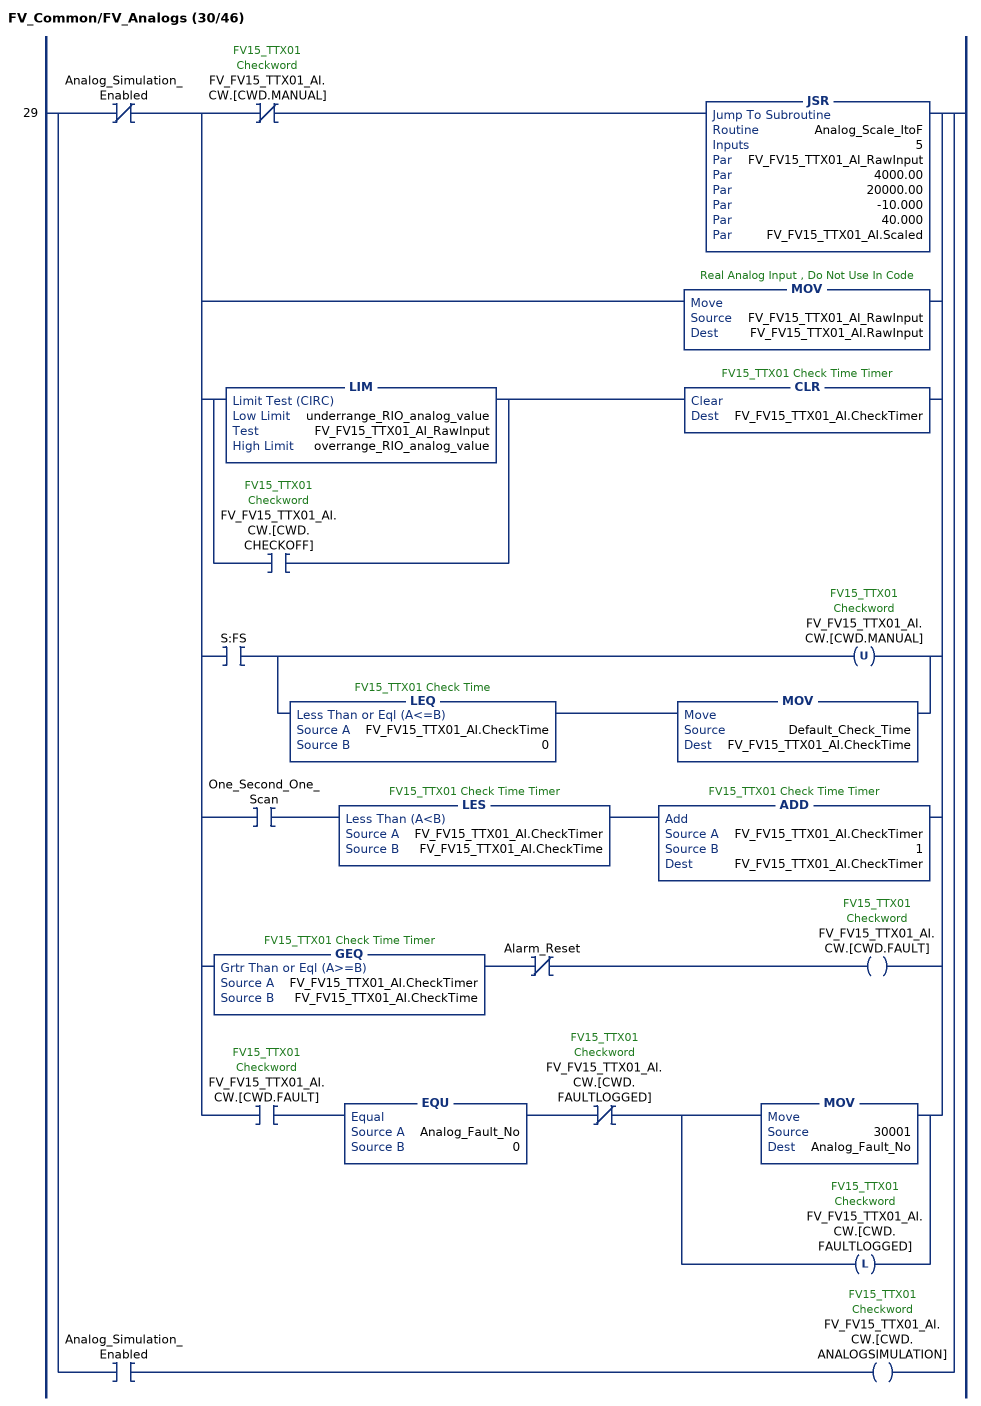
   29: [XIO(Analog_Simulation_Enabled) [XIO(FV_FV15_TTX01_AI.CW.[CWD.MANUAL]) JSR(Analog_Scale_ItoF,5,FV_FV15_TTX01_AI_RawInput,4000.00,20000.00,-10.000,40.000,FV_FV15_TTX01_AI.Scaled) ,MOV(FV_FV15_TTX01_AI_RawInput,FV_FV15_TTX01_AI.RawInput) ,[LIM(underrange_RIO_analog_value,FV_FV15_TTX01_AI_RawInput,overrange_RIO_analog_value) ,XIC(FV_FV15_TTX01_AI.CW.[CWD.CHECKOFF]) ] CLR(FV_FV15_TTX01_AI.CheckTimer) ,XIC(S:FS) [OTU(FV_FV15_TTX01_AI.CW.[CWD.MANUAL]) ,LEQ(FV_FV15_TTX01_AI.CheckTime,0) MOV(Default_Check_Time,FV_FV15_TTX01_AI.CheckTime) ] ,XIC(One_Second_One_Scan) LES(FV_FV15_TTX01_AI.CheckTimer,FV_FV15_TTX01_AI.CheckTime) ADD(FV_FV15_TTX01_AI.CheckTimer,1,FV_FV15_TTX01_AI.CheckTimer) ,GEQ(FV_FV15_TTX01_AI.CheckTimer,FV_FV15_TTX01_AI.CheckTime) XIO(Alarm_Reset) OTE(FV_FV15_TTX01_AI.CW.[CWD.FAULT]) ,XIC(FV_FV15_TTX01_AI.CW.[CWD.FAULT]) EQU(Analog_Fault_No,0) XIO(FV_FV15_TTX01_AI.CW.[CWD.FAULTLOGGED]) [MOV(30001,Analog_Fault_No) ,OTL(FV_FV15_TTX01_AI.CW.[CWD.FAULTLOGGED]) ] ] ,XIC(Analog_Simulation_Enabled) OTE(FV_FV15_TTX01_AI.CW.[CWD.ANALOGSIMULATION]) ];
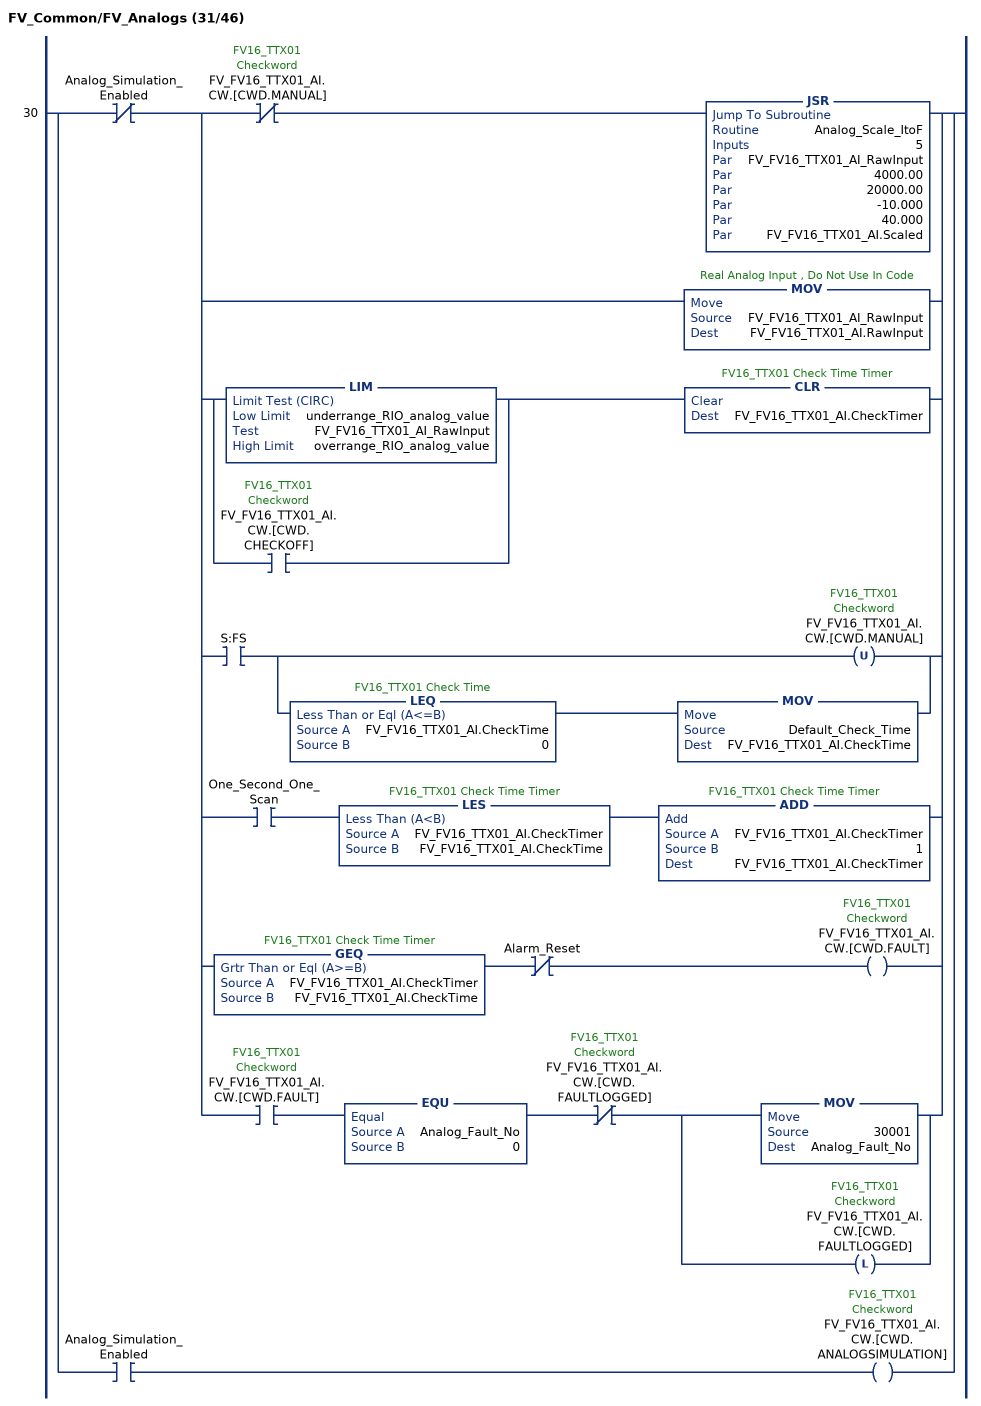
   30: [XIO(Analog_Simulation_Enabled) [XIO(FV_FV16_TTX01_AI.CW.[CWD.MANUAL]) JSR(Analog_Scale_ItoF,5,FV_FV16_TTX01_AI_RawInput,4000.00,20000.00,-10.000,40.000,FV_FV16_TTX01_AI.Scaled) ,MOV(FV_FV16_TTX01_AI_RawInput,FV_FV16_TTX01_AI.RawInput) ,[LIM(underrange_RIO_analog_value,FV_FV16_TTX01_AI_RawInput,overrange_RIO_analog_value) ,XIC(FV_FV16_TTX01_AI.CW.[CWD.CHECKOFF]) ] CLR(FV_FV16_TTX01_AI.CheckTimer) ,XIC(S:FS) [OTU(FV_FV16_TTX01_AI.CW.[CWD.MANUAL]) ,LEQ(FV_FV16_TTX01_AI.CheckTime,0) MOV(Default_Check_Time,FV_FV16_TTX01_AI.CheckTime) ] ,XIC(One_Second_One_Scan) LES(FV_FV16_TTX01_AI.CheckTimer,FV_FV16_TTX01_AI.CheckTime) ADD(FV_FV16_TTX01_AI.CheckTimer,1,FV_FV16_TTX01_AI.CheckTimer) ,GEQ(FV_FV16_TTX01_AI.CheckTimer,FV_FV16_TTX01_AI.CheckTime) XIO(Alarm_Reset) OTE(FV_FV16_TTX01_AI.CW.[CWD.FAULT]) ,XIC(FV_FV16_TTX01_AI.CW.[CWD.FAULT]) EQU(Analog_Fault_No,0) XIO(FV_FV16_TTX01_AI.CW.[CWD.FAULTLOGGED]) [MOV(30001,Analog_Fault_No) ,OTL(FV_FV16_TTX01_AI.CW.[CWD.FAULTLOGGED]) ] ] ,XIC(Analog_Simulation_Enabled) OTE(FV_FV16_TTX01_AI.CW.[CWD.ANALOGSIMULATION]) ];
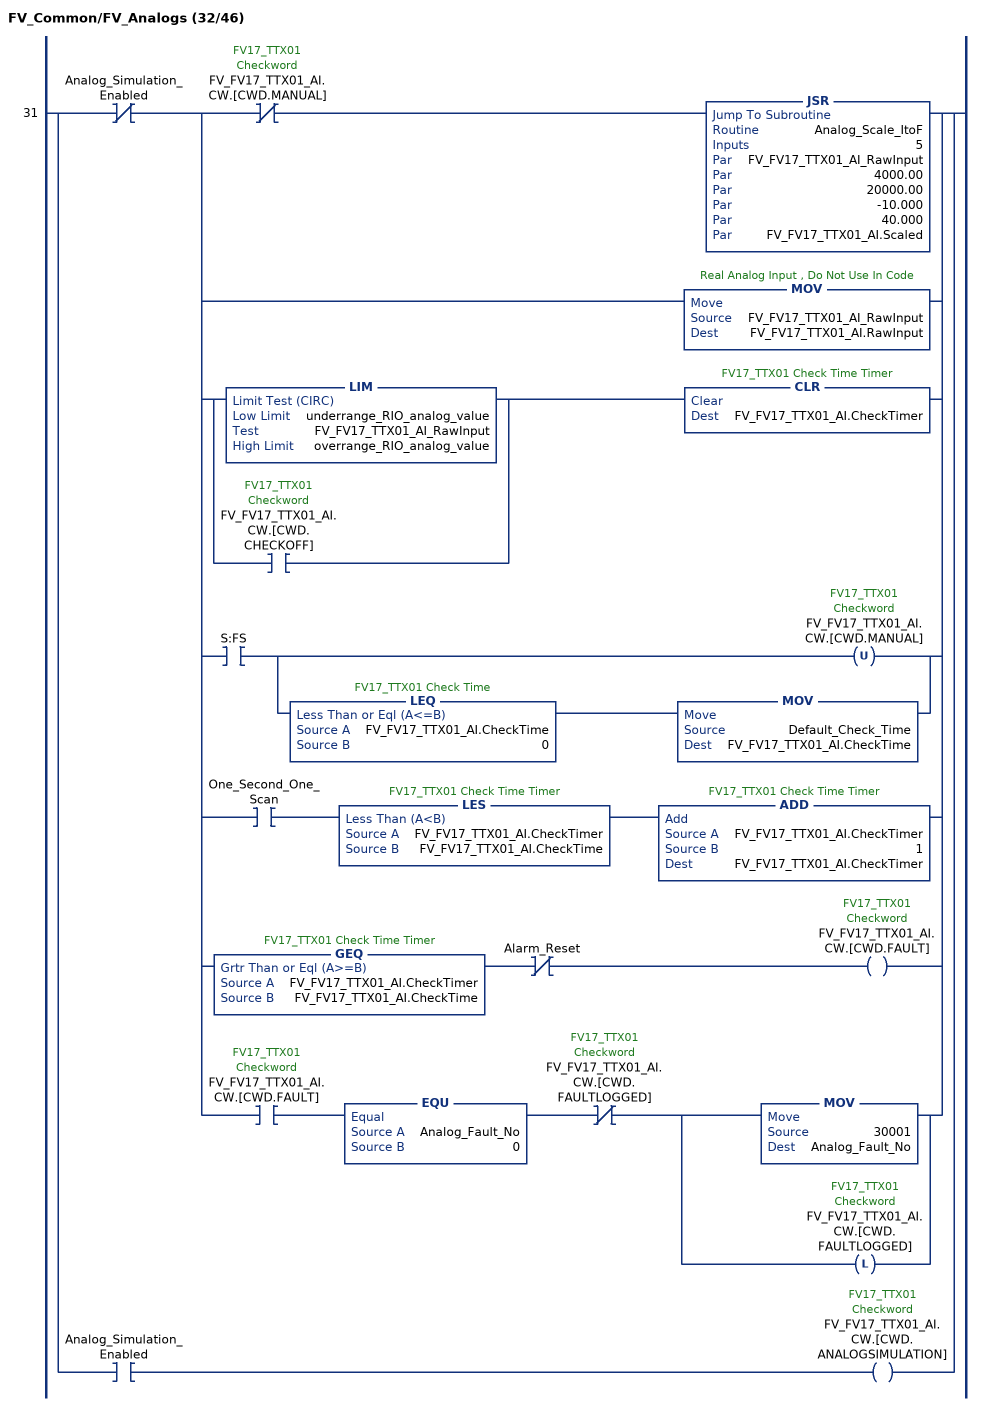
   31: [XIO(Analog_Simulation_Enabled) [XIO(FV_FV17_TTX01_AI.CW.[CWD.MANUAL]) JSR(Analog_Scale_ItoF,5,FV_FV17_TTX01_AI_RawInput,4000.00,20000.00,-10.000,40.000,FV_FV17_TTX01_AI.Scaled) ,MOV(FV_FV17_TTX01_AI_RawInput,FV_FV17_TTX01_AI.RawInput) ,[LIM(underrange_RIO_analog_value,FV_FV17_TTX01_AI_RawInput,overrange_RIO_analog_value) ,XIC(FV_FV17_TTX01_AI.CW.[CWD.CHECKOFF]) ] CLR(FV_FV17_TTX01_AI.CheckTimer) ,XIC(S:FS) [OTU(FV_FV17_TTX01_AI.CW.[CWD.MANUAL]) ,LEQ(FV_FV17_TTX01_AI.CheckTime,0) MOV(Default_Check_Time,FV_FV17_TTX01_AI.CheckTime) ] ,XIC(One_Second_One_Scan) LES(FV_FV17_TTX01_AI.CheckTimer,FV_FV17_TTX01_AI.CheckTime) ADD(FV_FV17_TTX01_AI.CheckTimer,1,FV_FV17_TTX01_AI.CheckTimer) ,GEQ(FV_FV17_TTX01_AI.CheckTimer,FV_FV17_TTX01_AI.CheckTime) XIO(Alarm_Reset) OTE(FV_FV17_TTX01_AI.CW.[CWD.FAULT]) ,XIC(FV_FV17_TTX01_AI.CW.[CWD.FAULT]) EQU(Analog_Fault_No,0) XIO(FV_FV17_TTX01_AI.CW.[CWD.FAULTLOGGED]) [MOV(30001,Analog_Fault_No) ,OTL(FV_FV17_TTX01_AI.CW.[CWD.FAULTLOGGED]) ] ] ,XIC(Analog_Simulation_Enabled) OTE(FV_FV17_TTX01_AI.CW.[CWD.ANALOGSIMULATION]) ];
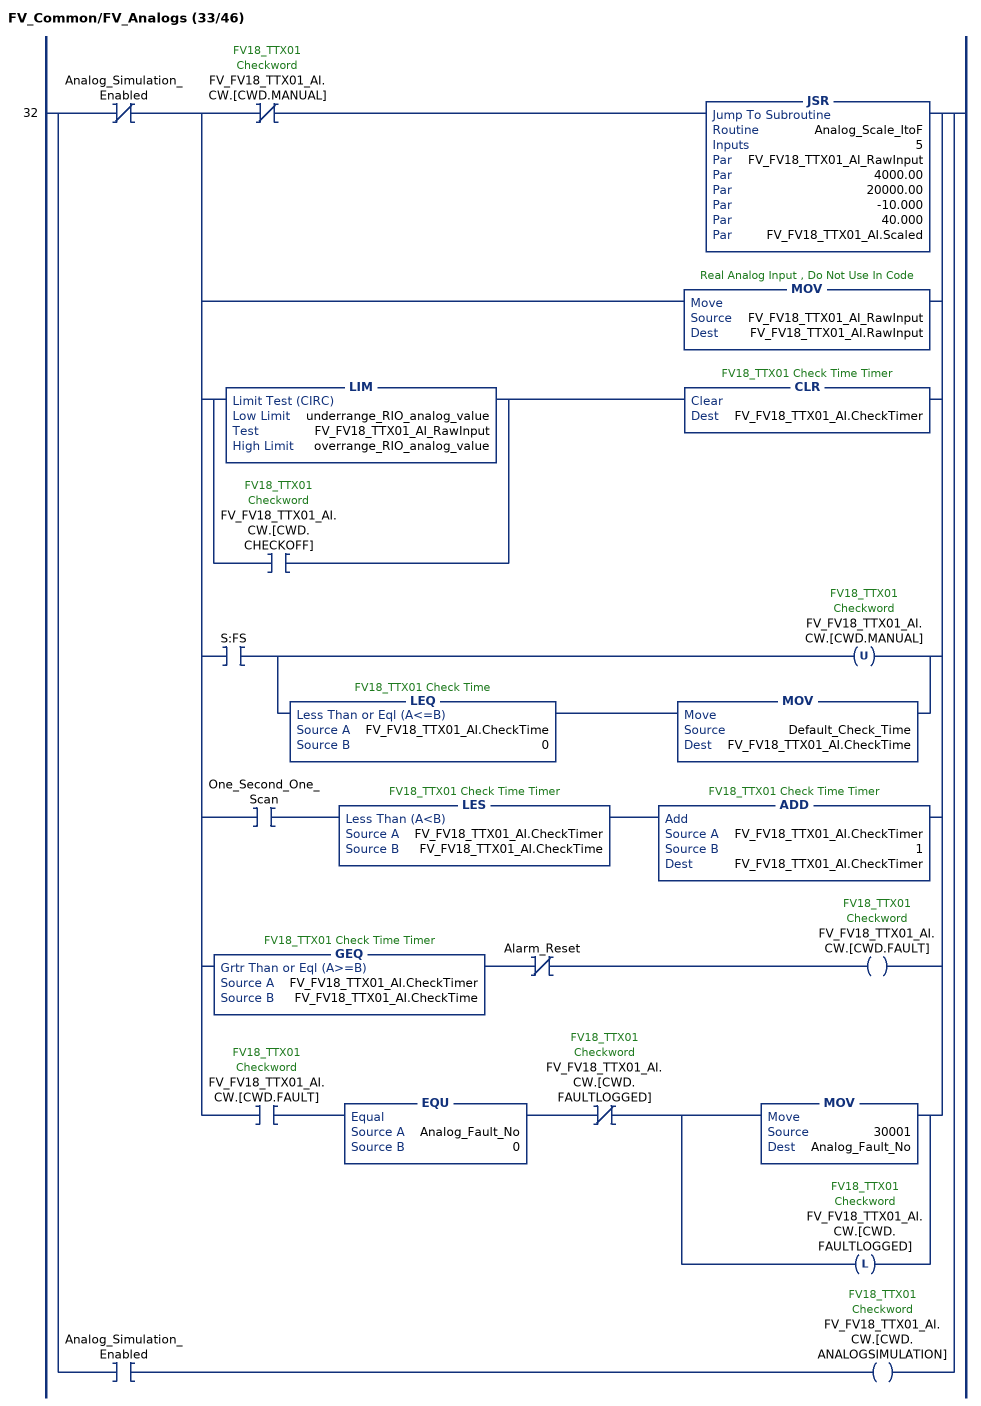
   32: [XIO(Analog_Simulation_Enabled) [XIO(FV_FV18_TTX01_AI.CW.[CWD.MANUAL]) JSR(Analog_Scale_ItoF,5,FV_FV18_TTX01_AI_RawInput,4000.00,20000.00,-10.000,40.000,FV_FV18_TTX01_AI.Scaled) ,MOV(FV_FV18_TTX01_AI_RawInput,FV_FV18_TTX01_AI.RawInput) ,[LIM(underrange_RIO_analog_value,FV_FV18_TTX01_AI_RawInput,overrange_RIO_analog_value) ,XIC(FV_FV18_TTX01_AI.CW.[CWD.CHECKOFF]) ] CLR(FV_FV18_TTX01_AI.CheckTimer) ,XIC(S:FS) [OTU(FV_FV18_TTX01_AI.CW.[CWD.MANUAL]) ,LEQ(FV_FV18_TTX01_AI.CheckTime,0) MOV(Default_Check_Time,FV_FV18_TTX01_AI.CheckTime) ] ,XIC(One_Second_One_Scan) LES(FV_FV18_TTX01_AI.CheckTimer,FV_FV18_TTX01_AI.CheckTime) ADD(FV_FV18_TTX01_AI.CheckTimer,1,FV_FV18_TTX01_AI.CheckTimer) ,GEQ(FV_FV18_TTX01_AI.CheckTimer,FV_FV18_TTX01_AI.CheckTime) XIO(Alarm_Reset) OTE(FV_FV18_TTX01_AI.CW.[CWD.FAULT]) ,XIC(FV_FV18_TTX01_AI.CW.[CWD.FAULT]) EQU(Analog_Fault_No,0) XIO(FV_FV18_TTX01_AI.CW.[CWD.FAULTLOGGED]) [MOV(30001,Analog_Fault_No) ,OTL(FV_FV18_TTX01_AI.CW.[CWD.FAULTLOGGED]) ] ] ,XIC(Analog_Simulation_Enabled) OTE(FV_FV18_TTX01_AI.CW.[CWD.ANALOGSIMULATION]) ];
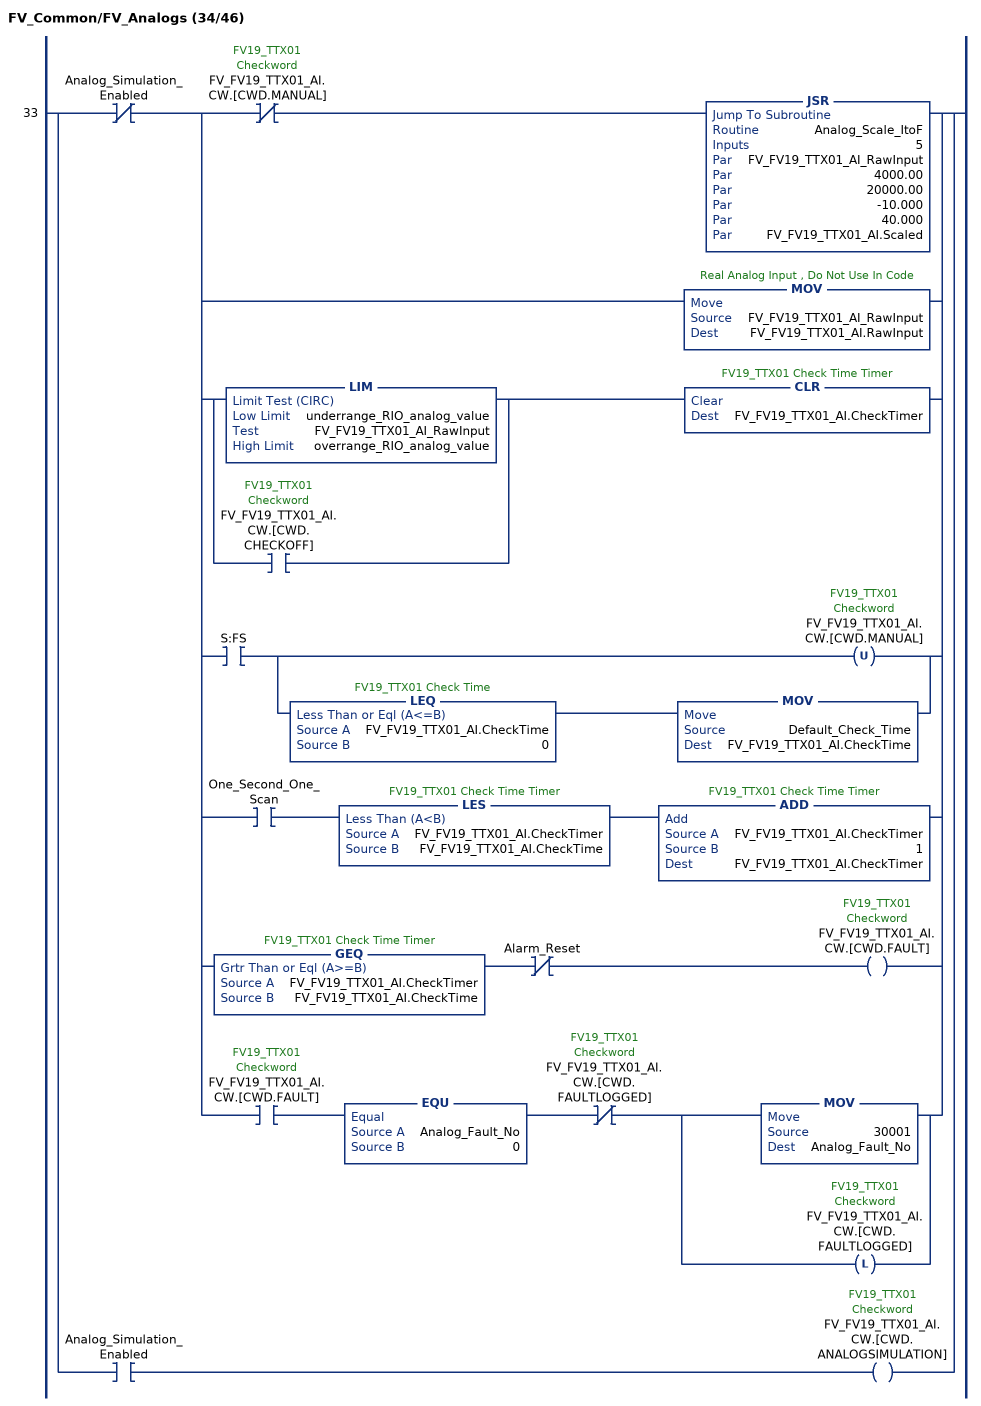
   33: [XIO(Analog_Simulation_Enabled) [XIO(FV_FV19_TTX01_AI.CW.[CWD.MANUAL]) JSR(Analog_Scale_ItoF,5,FV_FV19_TTX01_AI_RawInput,4000.00,20000.00,-10.000,40.000,FV_FV19_TTX01_AI.Scaled) ,MOV(FV_FV19_TTX01_AI_RawInput,FV_FV19_TTX01_AI.RawInput) ,[LIM(underrange_RIO_analog_value,FV_FV19_TTX01_AI_RawInput,overrange_RIO_analog_value) ,XIC(FV_FV19_TTX01_AI.CW.[CWD.CHECKOFF]) ] CLR(FV_FV19_TTX01_AI.CheckTimer) ,XIC(S:FS) [OTU(FV_FV19_TTX01_AI.CW.[CWD.MANUAL]) ,LEQ(FV_FV19_TTX01_AI.CheckTime,0) MOV(Default_Check_Time,FV_FV19_TTX01_AI.CheckTime) ] ,XIC(One_Second_One_Scan) LES(FV_FV19_TTX01_AI.CheckTimer,FV_FV19_TTX01_AI.CheckTime) ADD(FV_FV19_TTX01_AI.CheckTimer,1,FV_FV19_TTX01_AI.CheckTimer) ,GEQ(FV_FV19_TTX01_AI.CheckTimer,FV_FV19_TTX01_AI.CheckTime) XIO(Alarm_Reset) OTE(FV_FV19_TTX01_AI.CW.[CWD.FAULT]) ,XIC(FV_FV19_TTX01_AI.CW.[CWD.FAULT]) EQU(Analog_Fault_No,0) XIO(FV_FV19_TTX01_AI.CW.[CWD.FAULTLOGGED]) [MOV(30001,Analog_Fault_No) ,OTL(FV_FV19_TTX01_AI.CW.[CWD.FAULTLOGGED]) ] ] ,XIC(Analog_Simulation_Enabled) OTE(FV_FV19_TTX01_AI.CW.[CWD.ANALOGSIMULATION]) ];
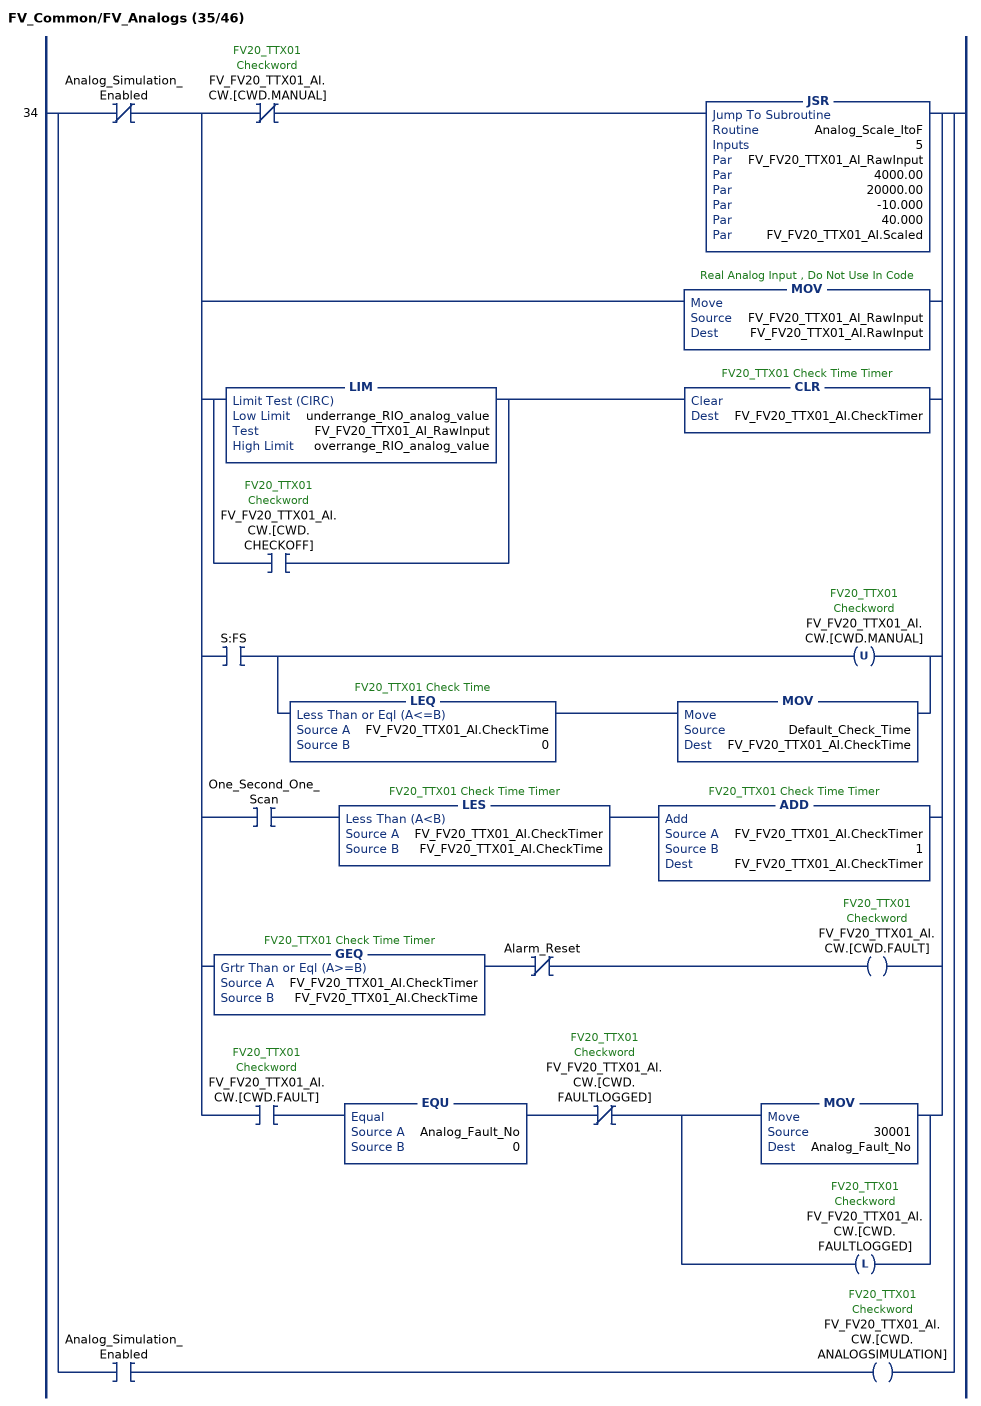
   34: [XIO(Analog_Simulation_Enabled) [XIO(FV_FV20_TTX01_AI.CW.[CWD.MANUAL]) JSR(Analog_Scale_ItoF,5,FV_FV20_TTX01_AI_RawInput,4000.00,20000.00,-10.000,40.000,FV_FV20_TTX01_AI.Scaled) ,MOV(FV_FV20_TTX01_AI_RawInput,FV_FV20_TTX01_AI.RawInput) ,[LIM(underrange_RIO_analog_value,FV_FV20_TTX01_AI_RawInput,overrange_RIO_analog_value) ,XIC(FV_FV20_TTX01_AI.CW.[CWD.CHECKOFF]) ] CLR(FV_FV20_TTX01_AI.CheckTimer) ,XIC(S:FS) [OTU(FV_FV20_TTX01_AI.CW.[CWD.MANUAL]) ,LEQ(FV_FV20_TTX01_AI.CheckTime,0) MOV(Default_Check_Time,FV_FV20_TTX01_AI.CheckTime) ] ,XIC(One_Second_One_Scan) LES(FV_FV20_TTX01_AI.CheckTimer,FV_FV20_TTX01_AI.CheckTime) ADD(FV_FV20_TTX01_AI.CheckTimer,1,FV_FV20_TTX01_AI.CheckTimer) ,GEQ(FV_FV20_TTX01_AI.CheckTimer,FV_FV20_TTX01_AI.CheckTime) XIO(Alarm_Reset) OTE(FV_FV20_TTX01_AI.CW.[CWD.FAULT]) ,XIC(FV_FV20_TTX01_AI.CW.[CWD.FAULT]) EQU(Analog_Fault_No,0) XIO(FV_FV20_TTX01_AI.CW.[CWD.FAULTLOGGED]) [MOV(30001,Analog_Fault_No) ,OTL(FV_FV20_TTX01_AI.CW.[CWD.FAULTLOGGED]) ] ] ,XIC(Analog_Simulation_Enabled) OTE(FV_FV20_TTX01_AI.CW.[CWD.ANALOGSIMULATION]) ];
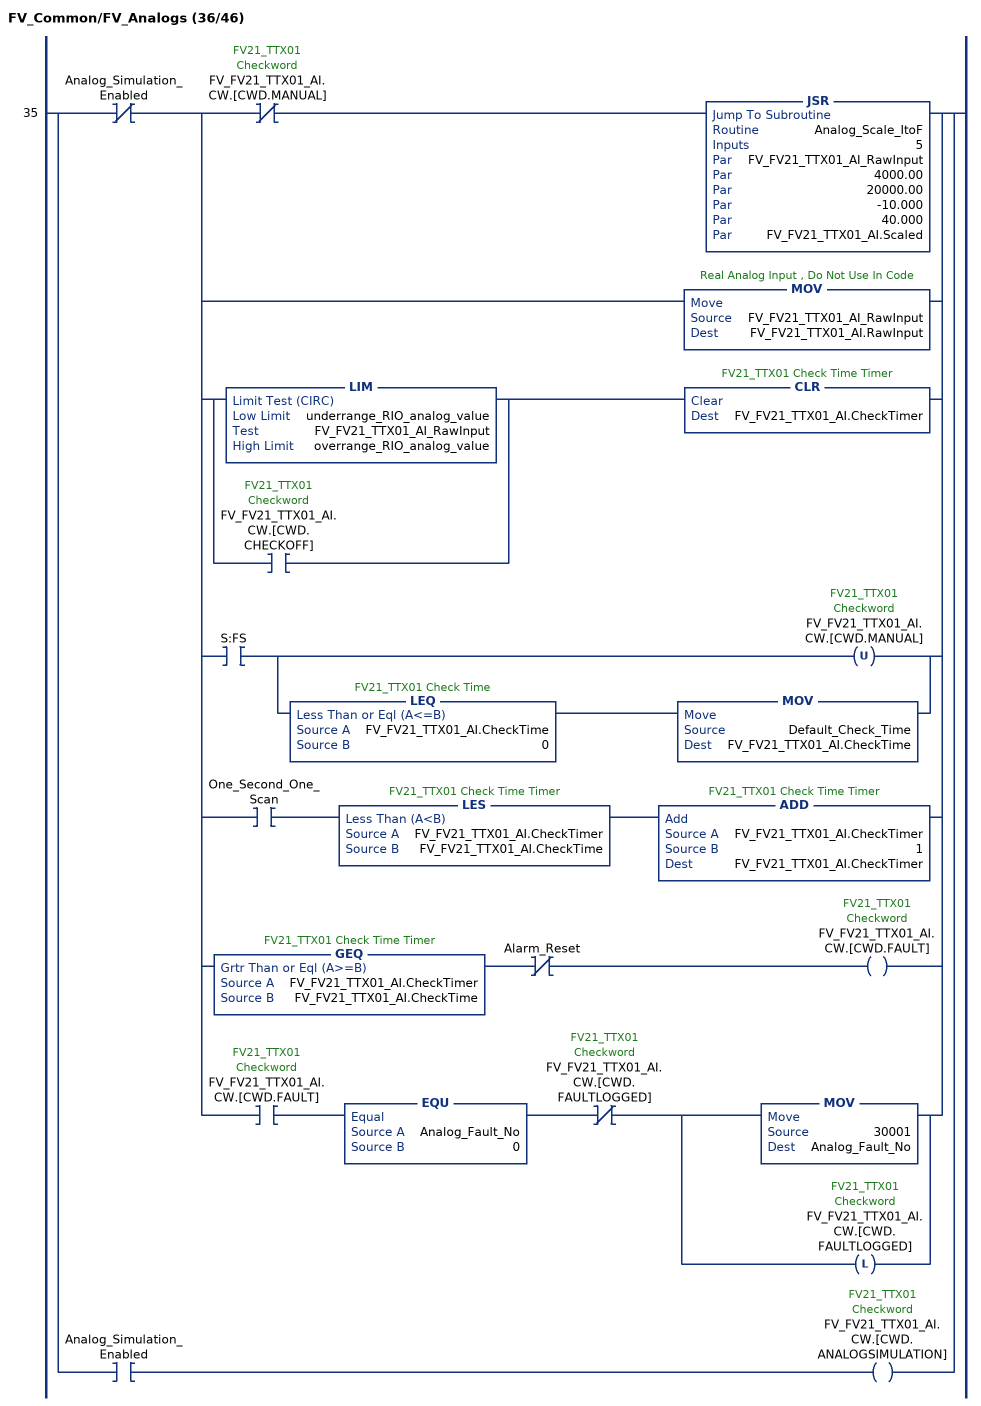
   35: [XIO(Analog_Simulation_Enabled) [XIO(FV_FV21_TTX01_AI.CW.[CWD.MANUAL]) JSR(Analog_Scale_ItoF,5,FV_FV21_TTX01_AI_RawInput,4000.00,20000.00,-10.000,40.000,FV_FV21_TTX01_AI.Scaled) ,MOV(FV_FV21_TTX01_AI_RawInput,FV_FV21_TTX01_AI.RawInput) ,[LIM(underrange_RIO_analog_value,FV_FV21_TTX01_AI_RawInput,overrange_RIO_analog_value) ,XIC(FV_FV21_TTX01_AI.CW.[CWD.CHECKOFF]) ] CLR(FV_FV21_TTX01_AI.CheckTimer) ,XIC(S:FS) [OTU(FV_FV21_TTX01_AI.CW.[CWD.MANUAL]) ,LEQ(FV_FV21_TTX01_AI.CheckTime,0) MOV(Default_Check_Time,FV_FV21_TTX01_AI.CheckTime) ] ,XIC(One_Second_One_Scan) LES(FV_FV21_TTX01_AI.CheckTimer,FV_FV21_TTX01_AI.CheckTime) ADD(FV_FV21_TTX01_AI.CheckTimer,1,FV_FV21_TTX01_AI.CheckTimer) ,GEQ(FV_FV21_TTX01_AI.CheckTimer,FV_FV21_TTX01_AI.CheckTime) XIO(Alarm_Reset) OTE(FV_FV21_TTX01_AI.CW.[CWD.FAULT]) ,XIC(FV_FV21_TTX01_AI.CW.[CWD.FAULT]) EQU(Analog_Fault_No,0) XIO(FV_FV21_TTX01_AI.CW.[CWD.FAULTLOGGED]) [MOV(30001,Analog_Fault_No) ,OTL(FV_FV21_TTX01_AI.CW.[CWD.FAULTLOGGED]) ] ] ,XIC(Analog_Simulation_Enabled) OTE(FV_FV21_TTX01_AI.CW.[CWD.ANALOGSIMULATION]) ];
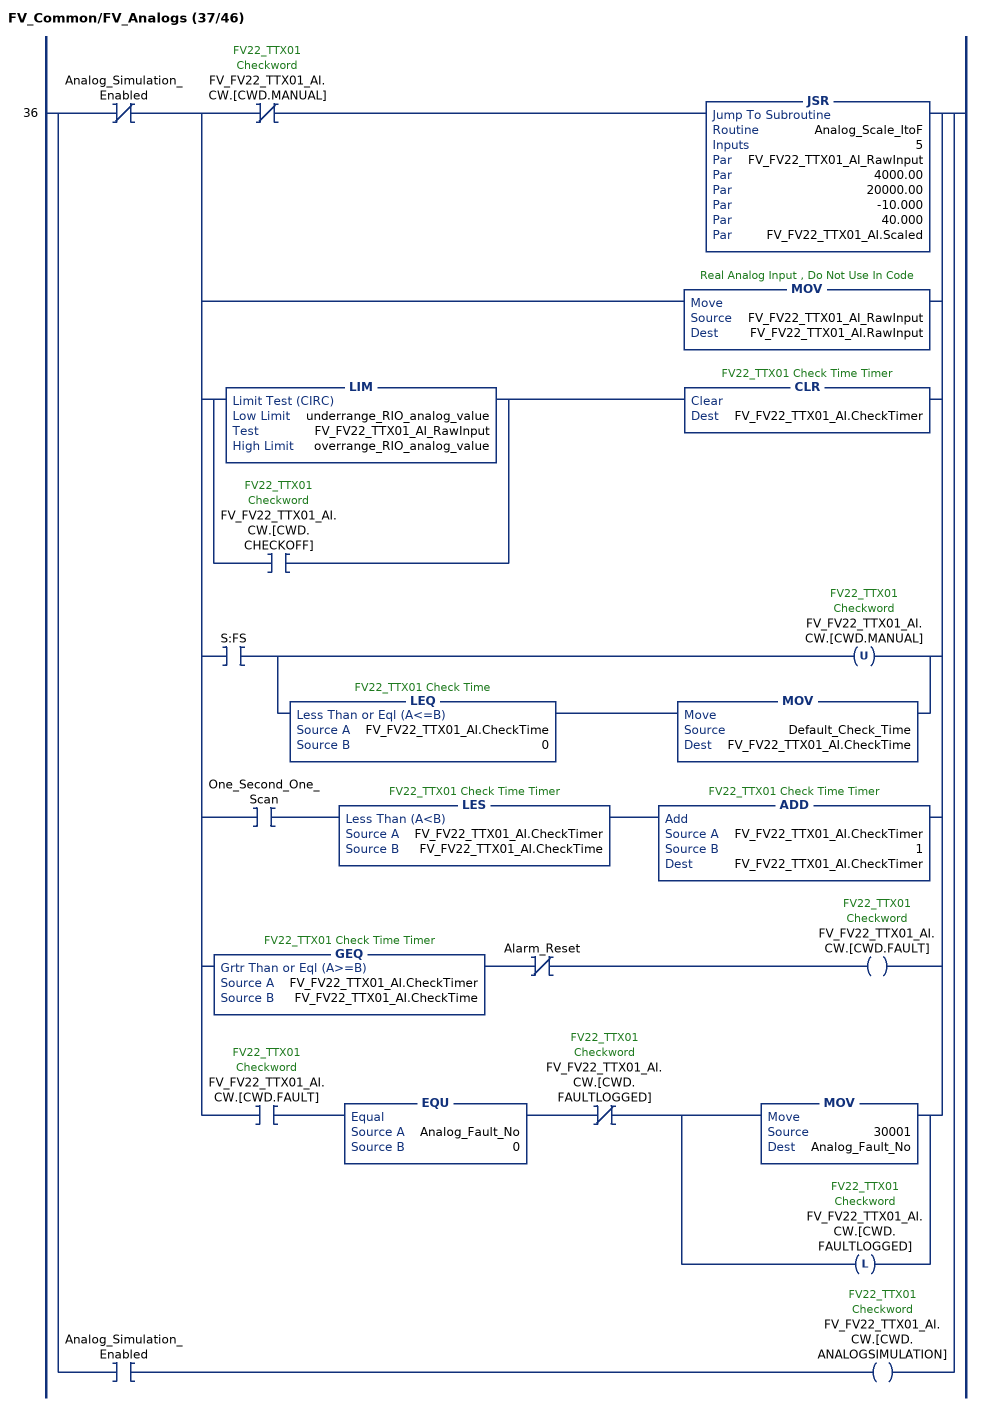
   36: [XIO(Analog_Simulation_Enabled) [XIO(FV_FV22_TTX01_AI.CW.[CWD.MANUAL]) JSR(Analog_Scale_ItoF,5,FV_FV22_TTX01_AI_RawInput,4000.00,20000.00,-10.000,40.000,FV_FV22_TTX01_AI.Scaled) ,MOV(FV_FV22_TTX01_AI_RawInput,FV_FV22_TTX01_AI.RawInput) ,[LIM(underrange_RIO_analog_value,FV_FV22_TTX01_AI_RawInput,overrange_RIO_analog_value) ,XIC(FV_FV22_TTX01_AI.CW.[CWD.CHECKOFF]) ] CLR(FV_FV22_TTX01_AI.CheckTimer) ,XIC(S:FS) [OTU(FV_FV22_TTX01_AI.CW.[CWD.MANUAL]) ,LEQ(FV_FV22_TTX01_AI.CheckTime,0) MOV(Default_Check_Time,FV_FV22_TTX01_AI.CheckTime) ] ,XIC(One_Second_One_Scan) LES(FV_FV22_TTX01_AI.CheckTimer,FV_FV22_TTX01_AI.CheckTime) ADD(FV_FV22_TTX01_AI.CheckTimer,1,FV_FV22_TTX01_AI.CheckTimer) ,GEQ(FV_FV22_TTX01_AI.CheckTimer,FV_FV22_TTX01_AI.CheckTime) XIO(Alarm_Reset) OTE(FV_FV22_TTX01_AI.CW.[CWD.FAULT]) ,XIC(FV_FV22_TTX01_AI.CW.[CWD.FAULT]) EQU(Analog_Fault_No,0) XIO(FV_FV22_TTX01_AI.CW.[CWD.FAULTLOGGED]) [MOV(30001,Analog_Fault_No) ,OTL(FV_FV22_TTX01_AI.CW.[CWD.FAULTLOGGED]) ] ] ,XIC(Analog_Simulation_Enabled) OTE(FV_FV22_TTX01_AI.CW.[CWD.ANALOGSIMULATION]) ];